      ProcessValue <- "MotorControl_Velocity_Velocity"
   Rectangle "Rectángulo_20" at 35,182 size 15x41
      Visibility <- "MotorControl_Velocity_Execute"
   Rectangle "Rectángulo_21" at 51,182 size 15x41
      Visibility <- "MotorControl_Velocity_Error"
   Rectangle "Rectángulo_22" at 19,182 size 15x41
      Visibility <- "MotorControl_Velocity_invelocity"
   TextField "Campo de texto_1" at 395,189 size 115x29; Text 'Velocidad / Velocity'
   IOField "Campo ES_7" at 524,13 size 142x40; FormatPattern s9999999999
      ProcessValue <- "2_PWMValve_Frecuency"
   TextField "Campo de texto_5" at 667,18 size 127x29; Text 'Frecuencia / Frequency'
   IOField "Campo ES_8" at 523,67 size 145x40; FormatPattern s99999
      ProcessValue <- "2_PWMValve_Duty_Cycle"
   TextField "Campo de texto_10" at 675,72 size 94x29; Text 'Trabajo / Duty'
   Rectangle "Rectángulo_18" at 575,117 size 15x41
      Visibility <- "2_PWMValve_Enable"
   Rectangle "Rectángulo_19" at 591,117 size 15x41
      Visibility <- "2_PWMValve_Busy"
   Rectangle "Rectángulo_38" at 559,117 size 15x41
      Visibility <- "2_PWMValve_Status"
   Button "Botón_9" at 610,184 size 145x40; TextOff 'MEM VELOC. / MEM SPEED'
      on Press: function_b14e0dd5("MotorControl_Velocity_Current", 0)
   TextField "Campo de texto_9" at 524,445 size 101x27; Text 'BATERIA / BATTERY'
   IOField "Campo ES_14" at 619,442 size 89x35; FormatPattern 99.9; Unit  Vdc
      ProcessValue <- "DataValues_BatteryVoltage"
   Button "Botón_14" at 534,442 size 35x35; TextOff 'M'
      on Press: ActivateScreen("Start", 0)
   IOField "Campo ES_15" at 711,442 size 82x35; FormatPattern 999.9; Unit  %
      ProcessValue <- "DataValues_BatteryCapacity"
   Button "Botón_18" at 582,442 size 35x35; TextOff 'M'
      on Press: ActivateScreen("Motor", 0)
   Button "Botón_1" at 7,442 size 80x35; TextOff 'GRAFICOS / GRAPHICS'
      on Press: ActivateScreen("Graphics", 0)
   Button "Botón_3" at 92,442 size 80x35; TextOff 'DATOS / DATA'
      on Press: ActivateScreen("Parameters", 0)
   Button "Botón_4" at 347,442 size 80x35; TextOff 'MANUALES / MANUALS'
      on Press: ActivateScreen("UserManual", 0)
   Button "Botón_5" at 432,442 size 80x35; TextOff 'ALARMAS / ALARMS'
      on Press: ActivateScreen("Alarms", 0)
   Button "Botón_12" at 177,442 size 80x35; TextOff 'PACIENTE / PATIENT'
      on Press: function_efd93a16("PatientData", 0, 0, 1, -1, 1)
   Button "Botón_19" at 262,442 size 80x35; TextOff 'RPM / BPM'
      on Press: function_efd93a16("RespirationRatios", 0, 0, 1, -1, 1)
   IOField "Campo ES_9" at 243,57 size 142x40; FormatPattern 9999
      ProcessValue <- "TurnAxis_Position"
   TextField "Campo de texto_11" at 396,62 size 100x29; Text 'Posición / Position'

PopupScreen "ControlMode" 600x300
   TextField "Campo de texto_2" at 107,59 size 238x39; Text 'Selección TIPO / Select TYPE'
   TextField "Campo de texto_1" at 204,5 size 192x30; Text 'MODO CONTROL / CONTROL MODE'
   SymbolicIOField "Campo ES simbólico_1" at 114,119 size 360x47; TextOff '0'; TextOn '1'; TextList "ControlMode"
      ProcessValue <- "OperatingParameters_ControlMode"
   Button "Botón_6" at 429,255 size 146x32; TextOff 'Salida / Exit'
      on Click: function_efd93a16("ControlMode", 0, 0, 0, -1, 1)
   IOField "Campo ES_8" at 23,255 size 242x32; FormatPattern 99999999999999999999
      ProcessValue <- "DateTime_LocalDateOut"

PopupScreen "Alarm" 400x300
   TextField "Campo de texto_1" at 41,95 size 315x91; Text 'ALARMA / ALARM'

PopupScreen "PatientData" 600x300
   TextField "Campo de texto_2" at 167,65 size 60x29; Text 'Sexo / Sex'
   TextField "Campo de texto_3" at 264,113 size 166x29; Text 'Volumen Tidal / Tidal Volume'
   TextField "Campo de texto_10" at 53,113 size 80x29; Text 'Altura / Height'
   IOField "Campo ES_6" at 138,110 size 110x35; FormatPattern 9.99; Unit m
      ProcessValue <- "PatientData_PatientHeight"
   IOField "Campo ES_11" at 432,110 size 110x35; FormatPattern 999.9; Unit ml
      ProcessValue <- "PatientData_TidalVolume"
   TextField "Campo de texto_1" at 198,8 size 204x30; Text 'DATOS PACIENTE / PATIENT DATA'
   SymbolicIOField "Campo ES simbólico_1" at 227,61 size 233x37; TextOn '1'; TextOff '0'; TextList "PatientSex"
      ProcessValue <- "PatientData_PatientType"
   Button "Botón_6" at 429,255 size 146x32; TextOff 'Salida / Exit'
      on Click: function_efd93a16("PatientData", 0, 0, 0, -1, 1)
   IOField "Campo ES_8" at 23,255 size 242x32; FormatPattern 99999999999999999999
      ProcessValue <- "DateTime_LocalDateOut"

PopupScreen "Pip" 600x300
   TextField "Campo de texto_2" at 242,90 size 46x29; Text 'PIP'
   IOField "Campo ES_8" at 389,87 size 75x35; Authorization "Operación"; FormatPattern 999
      ProcessValue <- "DataValues_PipValue"
   IOField "Campo ES_2" at 290,87 size 75x35; FormatPattern 999
      ProcessValue <- "OperatingParameters_PipMax"
   IOField "Campo ES_3" at 44,87 size 75x35; FormatPattern 999
      ProcessValue <- "OperatingParameters_PipSetpoint"
      Visibility <- "OperatingParameters_ControlMode"
   TextField "Campo de texto_5" at 34,44 size 128x29; Text 'CONSIGNA / SETPOINT'
   TextField "Campo de texto_6" at 300,44 size 55x29; Text 'MAX'
   TextField "Campo de texto_7" at 388,44 size 81x29; Text 'VALOR / VALUE'
   TextField "Campo de texto_8" at 496,44 size 56x29; Text 'MIN'
   IOField "Campo ES_7" at 485,87 size 75x35; FormatPattern 999
      ProcessValue <- "OperatingParameters_PipMin"
   IOField "Campo ES_1" at 290,141 size 75x35; FormatPattern 999
      ProcessValue <- "ProcessData_PpipSetpointAlarmHI"
   IOField "Campo ES_4" at 485,141 size 75x35; FormatPattern 999
      ProcessValue <- "ProcessData_PipSetpointAlarmLOW"
   IOField "Campo ES_5" at 290,195 size 75x35; FormatPattern 999
      ProcessValue <- "ProcessData_PipSetpointPreAlarmHI"
   IOField "Campo ES_6" at 485,195 size 75x35; FormatPattern 999
      ProcessValue <- "ProcessData_PipSetpointPreAlarmLOW"
   TextField "Campo de texto_1" at 155,144 size 134x29; Text 'PIP Alarma / PIP Alarm'
   TextField "Campo de texto_3" at 131,196 size 158x29; Text 'PIP PreAlarm'
   TextField "Campo de texto_4" at 187,8 size 226x30; Text 'PARAMETROS PEEP / PIP PARAMETERS'
   Button "Botón_6" at 429,255 size 146x32; TextOff 'Salida / Exit'
      on Click: function_efd93a16("Pip", 0, 0, 0, -1, 1)
   IOField "Campo ES_9" at 23,255 size 242x32; FormatPattern 99999999999999999999
      ProcessValue <- "DateTime_LocalDateOut"
   GraphicIOField "PlotLight_Round_GN_1" at 369,105 size 17x17; PictureOff "gris"; PictureOn "amarillo"
      ProcessValue <- "AlarmsRaw_PipDisplayPreAlarmHI"
   GraphicIOField "PlotLight_Round_GN_2" at 466,105 size 17x17; PictureOff "gris"; PictureOn "rojo"
      ProcessValue <- "AlarmsRaw_PipDisplayAlarmLOW"
   GraphicIOField "PlotLight_Round_GN_3" at 369,87 size 17x17; PictureOff "gris"; PictureOn "rojo"
      ProcessValue <- "AlarmsRaw_PipDisplayAlarmHI"
   GraphicIOField "PlotLight_Round_GN_4" at 466,87 size 17x17; PictureOff "gris"; PictureOn "amarillo"
      ProcessValue <- "AlarmsRaw_PipDisplayPreAlarmLOW"

PopupScreen "Plateau" 600x300
   TextField "Campo de texto_2" at 193,89 size 92x29; Text 'Plateau'
   IOField "Campo ES_8" at 389,87 size 75x35; Authorization "Operación"; FormatPattern 999
      ProcessValue <- "DataValues_PlateauValue"
   IOField "Campo ES_2" at 290,87 size 75x35; FormatPattern 999
      ProcessValue <- "OperatingParameters_PlateauMax"
   TextField "Campo de texto_5" at 34,44 size 128x29; Text 'CONSIGNA / SETPOINT'
   TextField "Campo de texto_6" at 300,44 size 55x29; Text 'MAX'
   TextField "Campo de texto_7" at 387,44 size 81x29; Text 'VALOR / VALUE'
   TextField "Campo de texto_8" at 496,44 size 56x29; Text 'MIN'
   IOField "Campo ES_7" at 485,87 size 75x35; FormatPattern 999
      ProcessValue <- "OperatingParameters_PlateauMin"
   IOField "Campo ES_1" at 290,141 size 75x35; FormatPattern 999
      ProcessValue <- "ProcessData_PlateauSetpointAlarmHI"
   IOField "Campo ES_4" at 485,141 size 75x35; FormatPattern 999
      ProcessValue <- "ProcessData_PlateaukSetpointAlarmLOW"
   IOField "Campo ES_5" at 290,195 size 75x35; FormatPattern 999
      ProcessValue <- "ProcessData_PlateauSetpointPreAlarmHI"
   IOField "Campo ES_6" at 485,195 size 75x35; FormatPattern 999
      ProcessValue <- "ProcessData_PlateauSetpointPreAlarmLOW"
   TextField "Campo de texto_1" at 119,144 size 166x29; Text 'Plateau Alarm'
   TextField "Campo de texto_3" at 81,198 size 204x29; Text 'Plateau PreAlarm'
   TextField "Campo de texto_4" at 165,7 size 271x30; Text 'PARAMETROS PLATEAU / PLATEAU PARAMETERS'
   Button "Botón_6" at 429,255 size 146x32; TextOff 'Salida / Exit'
      on Click: function_efd93a16("Plateau", 0, 0, 0, -1, 1)
   IOField "Campo ES_9" at 23,255 size 242x32; FormatPattern 99999999999999999999
      ProcessValue <- "DateTime_LocalDateOut"
   GraphicIOField "PlotLight_Round_GN_1" at 368,106 size 17x17; PictureOff "gris"; PictureOn "amarillo"
      ProcessValue <- "AlarmsRaw_PlateauDisplayPreAlarmHI"
   GraphicIOField "PlotLight_Round_GN_7" at 465,106 size 17x17; PictureOff "gris"; PictureOn "rojo"
      ProcessValue <- "AlarmsRaw_PlateauDisplayAlarmLOW"
   GraphicIOField "PlotLight_Round_GN_13" at 368,88 size 17x17; PictureOff "gris"; PictureOn "rojo"
      ProcessValue <- "AlarmsRaw_PlateauDisplayAlarmHI"
   GraphicIOField "PlotLight_Round_GN_19" at 465,88 size 17x17; PictureOff "gris"; PictureOn "amarillo"
      ProcessValue <- "AlarmsRaw_PlateauDisplayPreAlarmLOW"

PopupScreen "Peep" 600x300
   TextField "Campo de texto_2" at 225,88 size 60x29; Text 'Peep'
   IOField "Campo ES_8" at 391,87 size 75x35; Authorization "Operación"; FormatPattern 999
      ProcessValue <- "DataValues_PeepValue"
   IOField "Campo ES_2" at 290,87 size 75x35; FormatPattern 999
      ProcessValue <- "OperatingParameters_PeepMax"
   IOField "Campo ES_3" at 44,87 size 75x35; FormatPattern 999
      ProcessValue <- "OperatingParameters_PeepSetpoint"
      Visibility <- "OperatingParameters_ControlMode"
   TextField "Campo de texto_5" at 34,44 size 128x29; Text 'CONSIGNA / SETPOINT'
   TextField "Campo de texto_6" at 300,44 size 55x29; Text 'MAX'
   TextField "Campo de texto_7" at 389,44 size 81x29; Text 'VALOR / VALUE'
   TextField "Campo de texto_8" at 496,44 size 56x29; Text 'MIN'
   IOField "Campo ES_7" at 485,87 size 75x35; FormatPattern 999
      ProcessValue <- "OperatingParameters_PeepMin"
   IOField "Campo ES_1" at 290,141 size 75x35; FormatPattern 999
      ProcessValue <- "ProcessData_PeepSetpointAlarmHI"
   IOField "Campo ES_4" at 485,141 size 75x35; FormatPattern 999
      ProcessValue <- "ProcessData_PeepSetpointAlarmLOW"
   IOField "Campo ES_5" at 290,195 size 75x35; FormatPattern 999
      ProcessValue <- "ProcessData_PeepSetpointPreAlarmHI"
   IOField "Campo ES_6" at 485,195 size 75x35; FormatPattern 999
      ProcessValue <- "ProcessData_PeepSetpointPreAlarmLOW"
   TextField "Campo de texto_1" at 141,143 size 148x29; Text 'Peep Alarma / Peep Alarm'
   TextField "Campo de texto_3" at 103,197 size 186x29; Text 'Peep PreAlarma / Peep PreAlarm'
   TextField "Campo de texto_4" at 187,8 size 226x30; Text 'PARAMETROS PEEP / PEEP PARAMETERS'
   Button "Botón_6" at 429,255 size 146x32; TextOff 'Salida / Exit'
      on Click: function_efd93a16("Peep", 0, 0, 0, -1, 1)
   IOField "Campo ES_9" at 23,255 size 242x32; FormatPattern 99999999999999999999
      ProcessValue <- "DateTime_LocalDateOut"
   GraphicIOField "PlotLight_Round_GN_2" at 370,104 size 17x17; PictureOff "gris"; PictureOn "amarillo"
      ProcessValue <- "AlarmsRaw_PeepDisplayPreAlarmHI"
   GraphicIOField "PlotLight_Round_GN_8" at 467,104 size 17x17; PictureOff "gris"; PictureOn "rojo"
      ProcessValue <- "AlarmsRaw_PeepDisplayAlarmLOW"
   GraphicIOField "PlotLight_Round_GN_14" at 370,86 size 17x17; PictureOff "gris"; PictureOn "rojo"
      ProcessValue <- "AlarmsRaw_PeepDisplayAlarmHI"
   GraphicIOField "PlotLight_Round_GN_20" at 467,86 size 17x17; PictureOff "gris"; PictureOn "amarillo"
      ProcessValue <- "AlarmsRaw_PeepDisplayPreAlarmLOW"

PopupScreen "Frecuency" 600x300
   TextField "Campo de texto_2" at 161,89 size 127x29; Text 'Frecuencia / Frequency'
   IOField "Campo ES_8" at 388,87 size 75x35; Authorization "Operación"; FormatPattern 999
      ProcessValue <- "DataValues_FrequencyValue"
   IOField "Campo ES_2" at 290,87 size 75x35; FormatPattern 999
      ProcessValue <- "OperatingParameters_FrequencyMax"
   IOField "Campo ES_3" at 44,87 size 75x35; FormatPattern 999
      ProcessValue <- "OperatingParameters_FrequencySetpoint"
   TextField "Campo de texto_5" at 34,44 size 128x29; Text 'CONSIGNA / SETPOINT'
   TextField "Campo de texto_6" at 300,44 size 55x29; Text 'MAX'
   TextField "Campo de texto_7" at 387,44 size 81x29; Text 'VALOR / VALUE'
   TextField "Campo de texto_8" at 496,44 size 56x29; Text 'MIN'
   IOField "Campo ES_7" at 485,87 size 75x35; FormatPattern 999
      ProcessValue <- "OperatingParameters_FrequencyMin"
   IOField "Campo ES_1" at 290,141 size 75x35; FormatPattern 999
      ProcessValue <- "ProcessData_FrequencySetpointAlarmHI"
   IOField "Campo ES_4" at 485,141 size 75x35; FormatPattern 999
      ProcessValue <- "ProcessData_FrequencySetpointAlarmLOW"
   IOField "Campo ES_5" at 290,195 size 75x35; FormatPattern 999
      ProcessValue <- "ProcessData_FrequencySetpointPreAlarmHI"
   IOField "Campo ES_6" at 485,195 size 75x35; FormatPattern 999
      ProcessValue <- "ProcessData_FrequencySetpointPreAlarmLOW"
   TextField "Campo de texto_1" at 73,144 size 215x29; Text 'Frecuencia Alarma / Frequency Alarm'
   TextField "Campo de texto_3" at 56,197 size 233x29; Text 'FrecuenciaPreAlarm / Frequency PreAlarm'
   TextField "Campo de texto_4" at 143,5 size 315x30; Text 'PARAMETROS FRECUENCIA / FREQUENCY PARAMETERS'
   Button "Botón_6" at 429,255 size 146x32; TextOff 'Salida / Exit'
      on Click: function_efd93a16("Frecuency", 0, 0, 0, -1, 1)
   IOField "Campo ES_9" at 23,255 size 242x32; FormatPattern 99999999999999999999
      ProcessValue <- "DateTime_LocalDateOut"
   GraphicIOField "PlotLight_Round_GN_3" at 369,105 size 17x17; PictureOff "gris"; PictureOn "amarillo"
      ProcessValue <- "AlarmsRaw_FrequencyDisplayPreAlarmHI"
   GraphicIOField "PlotLight_Round_GN_9" at 466,105 size 17x17; PictureOff "gris"; PictureOn "rojo"
      ProcessValue <- "AlarmsRaw_FrequencyDisplayAlarmLOW"
   GraphicIOField "PlotLight_Round_GN_15" at 369,87 size 17x17; PictureOff "gris"; PictureOn "rojo"
      ProcessValue <- "AlarmsRaw_FrequencyDisplayAlarmHI"
   GraphicIOField "PlotLight_Round_GN_21" at 466,87 size 17x17; PictureOff "gris"; PictureOn "amarillo"
      ProcessValue <- "AlarmsRaw_FrequencyDisplayPreAlarmLOW"

PopupScreen "TidalVolume" 600x300
   TextField "Campo de texto_2" at 123,90 size 166x29; Text 'Volumen Tidal / Tidal Volume'
   IOField "Campo ES_8" at 391,87 size 75x35; Authorization "Operación"; FormatPattern 999
      ProcessValue <- "DataValues_TidalVolumeValue"
   IOField "Campo ES_2" at 290,87 size 75x35; FormatPattern 999
      ProcessValue <- "OperatingParameters_TidalVolumenMax"
   IOField "Campo ES_3" at 44,87 size 75x35; FormatPattern 999
      ProcessValue <- "OperatingParameters_TidalVolumenSetpoint"
      Visibility <- "OperatingParameters_ControlMode"
   TextField "Campo de texto_5" at 34,44 size 128x29; Text 'CONSIGNA / SETPOINT'
   TextField "Campo de texto_6" at 300,44 size 55x29; Text 'MAX'
   TextField "Campo de texto_7" at 391,44 size 81x29; Text 'VALOR / VALUE'
   TextField "Campo de texto_8" at 496,44 size 56x29; Text 'MIN'
   IOField "Campo ES_7" at 485,87 size 75x35; FormatPattern 999
      ProcessValue <- "OperatingParameters_TidalVolumenMin"
   IOField "Campo ES_1" at 290,141 size 75x35; FormatPattern 999
      ProcessValue <- "ProcessData_TidalVolumeSetpointAlarmHI"
   IOField "Campo ES_4" at 485,141 size 75x35; FormatPattern 999
      ProcessValue <- "ProcessData_TidalVolumeSetpointAlarmLOW"
   IOField "Campo ES_5" at 290,195 size 75x35; FormatPattern 999
      ProcessValue <- "ProcessData_TidalVolumeSetpointPreAlarmHI"
   IOField "Campo ES_6" at 485,195 size 75x35; FormatPattern 999
      ProcessValue <- "ProcessData_TidalVolumeSetpointPreAlarmLOW"
   TextField "Campo de texto_1" at 35,143 size 254x29; Text 'Alarma Volumen Tidal / Tidal Volume Alarm'
   TextField "Campo de texto_3" at 0,197 size 290x29; Text 'PreAlarma volumen Tidal / Tidal Volume PreAlarm'
   TextField "Campo de texto_4" at 121,8 size 358x30; Text 'PARAMETROS VOLUMEN TIDAL / TIDAL VOLUME PARAMETERS'
   Button "Botón_6" at 429,255 size 146x32; TextOff 'Salida / Exit'
      on Click: function_efd93a16("TidalVolume", 0, 0, 0, -1, 1)
   IOField "Campo ES_9" at 23,255 size 242x32; FormatPattern 99999999999999999999
      ProcessValue <- "DateTime_LocalDateOut"
   GraphicIOField "PlotLight_Round_GN_4" at 370,105 size 17x17; PictureOff "gris"; PictureOn "amarillo"
      ProcessValue <- "AlarmsRaw_TidalVolumeDisplayPreAlarmHI"
   GraphicIOField "PlotLight_Round_GN_10" at 467,105 size 17x17; PictureOff "gris"; PictureOn "rojo"
      ProcessValue <- "AlarmsRaw_TidalVolumeDisplayAlarmLOW"
   GraphicIOField "PlotLight_Round_GN_16" at 370,87 size 17x17; PictureOff "gris"; PictureOn "rojo"
      ProcessValue <- "AlarmsRaw_TidalVolumeDisplayAlarmHI"
   GraphicIOField "PlotLight_Round_GN_22" at 467,87 size 17x17; PictureOff "gris"; PictureOn "amarillo"
      ProcessValue <- "AlarmsRaw_TidalVolumeDisplayPreAlarmLOW"

PopupScreen "VolumeMinute" 600x300
   TextField "Campo de texto_2" at 114,90 size 174x29; Text 'Vol. Minute / Minute Volume'
   IOField "Campo ES_8" at 388,87 size 75x35; Authorization "Operación"; FormatPattern 999
      ProcessValue <- "DataValues_MinumValue"
   IOField "Campo ES_2" at 290,87 size 75x35; FormatPattern 999
      ProcessValue <- "OperatingParameters_MinimumVolumeMax"
   IOField "Campo ES_3" at 44,87 size 75x35; FormatPattern 999
      Visibility <- "OperatingParameters_ControlMode"
      ProcessValue <- "OperatingParameters_MinimumVolumeSetpoint"
   TextField "Campo de texto_5" at 34,44 size 128x29; Text 'CONSIGNA / SETPOINT'
   TextField "Campo de texto_6" at 300,44 size 55x29; Text 'MAX'
   TextField "Campo de texto_7" at 390,44 size 81x29; Text 'VALOR / VALUE'
   TextField "Campo de texto_8" at 496,44 size 56x29; Text 'MIN'
   IOField "Campo ES_7" at 485,87 size 75x35; FormatPattern 999
      ProcessValue <- "OperatingParameters_MinimumVolumeMin"
   IOField "Campo ES_1" at 290,141 size 75x35; FormatPattern 999
      ProcessValue <- "ProcessData_VolumeMinSetpointAlarmHI"
   IOField "Campo ES_4" at 485,141 size 75x35; FormatPattern 999
      ProcessValue <- "ProcessData_VolumeMinSetpointPreAlarmLOW"
   IOField "Campo ES_5" at 290,195 size 75x35; FormatPattern 999
      ProcessValue <- "ProcessData_VolumeMinSetpointPreAlarmHI"
   IOField "Campo ES_6" at 485,195 size 75x35; FormatPattern 999
      ProcessValue <- "ProcessData_VolumeMinSetpointAlarmLOW"
   TextField "Campo de texto_1" at 20,143 size 269x29; Text 'Volumen/Minuto Alarm / Volume/Minute Alarm'
   TextField "Campo de texto_3" at 12,198 size 277x29; Text 'Volumen/Min. PreAlarm / Volume/Min. PreAlarm'
   TextField "Campo de texto_4" at 105,5 size 390x30; Text 'PARAMETROS VOLUMEN/MINUTO / VOLUME/MINUTE PARAMETERS'
   Button "Botón_6" at 429,255 size 146x32; TextOff 'Salida / Exit'
      on Click: function_efd93a16("VolumeMinute", 0, 0, 0, -1, 1)
   IOField "Campo ES_9" at 23,255 size 242x32; FormatPattern 99999999999999999999
      ProcessValue <- "DateTime_LocalDateOut"
   GraphicIOField "PlotLight_Round_GN_5" at 368,87 size 17x17; PictureOff "gris"; PictureOn "rojo"
      ProcessValue <- "AlarmsRaw_VolumeMinuteDisplayAlarmHI"
   GraphicIOField "PlotLight_Round_GN_11" at 465,105 size 17x17; PictureOff "gris"; PictureOn "rojo"
      ProcessValue <- "AlarmsRaw_VolumeMinuteDisplayAlarmLOW"
   GraphicIOField "PlotLight_Round_GN_17" at 368,105 size 17x17; PictureOff "gris"; PictureOn "amarillo"
      ProcessValue <- "AlarmsRaw_VolumeMinuteDisplayPreAlarmHI"
   GraphicIOField "PlotLight_Round_GN_23" at 465,87 size 17x17; PictureOff "gris"; PictureOn "amarillo"
      ProcessValue <- "AlarmsRaw_VolumeMinuteDisplayPreAlarmLOW"

PopupScreen "Trigger" 600x300
   TextField "Campo de texto_2" at 199,88 size 87x29; Text 'Trigger'
   IOField "Campo ES_8" at 388,87 size 75x35; Authorization "Operación"; FormatPattern 999
      ProcessValue <- "DataValues_Trigger"
   IOField "Campo ES_2" at 290,87 size 75x35; FormatPattern 999
      ProcessValue <- "OperatingParameters_TriggerMax"
   IOField "Campo ES_3" at 44,87 size 75x35; FormatPattern 999
      ProcessValue <- "OperatingParameters_TriggerSetpoint"
   TextField "Campo de texto_5" at 34,44 size 128x29; Text 'CONSIGNA / SETPOINT'
   TextField "Campo de texto_6" at 300,44 size 55x29; Text 'MAX'
   TextField "Campo de texto_7" at 387,44 size 81x29; Text 'VALOR / VALUE'
   TextField "Campo de texto_8" at 496,44 size 56x29; Text 'MIN'
   IOField "Campo ES_7" at 485,87 size 75x35; FormatPattern 999
      ProcessValue <- "OperatingParameters_TriggerMin"
   IOField "Campo ES_1" at 290,141 size 75x35; FormatPattern 999
      ProcessValue <- "ProcessData_TriggerVolumeSetpointAlarmHI"
   IOField "Campo ES_4" at 485,141 size 75x35; FormatPattern 999
      ProcessValue <- "ProcessData_TriggerVolumeSetpointAlarmLOW"
   IOField "Campo ES_5" at 290,195 size 75x35; FormatPattern 999
      ProcessValue <- "ProcessData_TriggeVolumeSetpointPreAlarmHI"
   IOField "Campo ES_6" at 485,195 size 75x35; FormatPattern 999
      ProcessValue <- "ProcessData_TriggerVolumeSetpointPreAlarmLOW"
   TextField "Campo de texto_1" at 125,143 size 161x29; Text 'Trigger Alarm'
   TextField "Campo de texto_3" at 87,197 size 199x29; Text 'Trigger PreAlarm'
   TextField "Campo de texto_4" at 164,8 size 273x30; Text 'PARAMETROS TRIGGER / TRIGGER PARAMETERS'
   Button "Botón_6" at 429,255 size 146x32; TextOff 'Salida / Exit'
      on Click: function_efd93a16("Trigger", 0, 0, 0, -1, 1)
   Button "Botón_7" at 396,141 size 61x35; TextOff 'Trigger'
      Visibility <- "Clock_1Hz"
   TextField "Campo de texto_9" at 396,196 size 61x35; Text 'OFF'
      Visibility <- "OperatingParameters_Trigger"
   TextField "Campo de texto_10" at 396,196 size 61x35; Text 'ON'
      Visibility <- "OperatingParameters_Trigger"
   Button "Botón_1" at 396,196 size 61x35; TextOn 'ON'; TextOff 'Text'
      on Click: InvertBit("OperatingParameters_Trigger")
      Appearance <- "OperatingParameters_Trigger"
   IOField "Campo ES_9" at 23,255 size 242x32; FormatPattern 99999999999999999999
      ProcessValue <- "DateTime_LocalDateOut"
   GraphicIOField "PlotLight_Round_GN_4" at 370,105 size 17x17; PictureOn "amarillo"; PictureOff "gris"
      ProcessValue <- "AlarmsRaw_TriggerDisplayPreAlarmHI"
   GraphicIOField "PlotLight_Round_GN_10" at 467,105 size 17x17; PictureOn "rojo"; PictureOff "gris"
      ProcessValue <- "AlarmsRaw_TriggerDisplayAlarmLOW"
   GraphicIOField "PlotLight_Round_GN_16" at 370,87 size 17x17; PictureOn "rojo"; PictureOff "gris"
      ProcessValue <- "AlarmsRaw_TriggerDisplayAlarmHI"
   GraphicIOField "PlotLight_Round_GN_22" at 467,87 size 17x17; PictureOn "amarillo"; PictureOff "gris"
      ProcessValue <- "AlarmsRaw_TriggerDisplayPreAlarmLOW"

PopupScreen "Enviroment" 600x300
   TextField "Campo de texto_2" at 30,82 size 124x29; Text 'Humidif. / Humidifier'
   IOField "Campo ES_3" at 246,192 size 75x35; FormatPattern 999
      ProcessValue <- "OperatingParameters_O2Setpoint"
   TextField "Campo de texto_4" at 140,5 size 320x30; Text 'PARAMETROS ENTORNO / ENVIROMENT PARAMETERS'
   Button "Botón_6" at 429,255 size 146x32; TextOff 'Salida / Exit'
      on Click: function_efd93a16("Enviroment", 0, 0, 0, -1, 1)
   Button "Botón_7" at 429,79 size 61x35; TextOff 'Hr'
      Visibility <- "Clock_1Hz"
   TextField "Campo de texto_9" at 502,79 size 61x35; Text 'OFF'
      Visibility <- "OperatingParameters_Trigger"
   TextField "Campo de texto_10" at 502,79 size 61x35; Text 'ON'
      Visibility <- "OperatingParameters_Trigger"
   Button "Botón_1" at 506,79 size 61x35; TextOn 'ON'; TextOff 'Text'
      on Click: InvertBit("OperatingParameters_Trigger")
      Appearance <- "OperatingParameters_Trigger"
   IOField "Campo ES_5" at 330,80 size 89x35; FormatPattern 9999999
      ProcessValue <- "OperatingParameters_HumidifiertElap"
   IOField "Campo ES_1" at 237,80 size 89x35; FormatPattern 9999999
      ProcessValue <- "OperatingParameters_HumidifierTimer"
   TextField "Campo de texto_1" at 38,196 size 142x29; Text 'Presión O2 / O2 Pressure'
   Button "Botón_2" at 429,192 size 61x35; TextOff 'O2'
      Visibility <- "Clock_1Hz"
   TextField "Campo de texto_3" at 502,192 size 61x35; Text 'OFF'
      Visibility <- "OperatingParameters_O2"
   TextField "Campo de texto_5" at 502,192 size 61x35; Text 'ON'
      Visibility <- "OperatingParameters_O2"
   Button "Botón_3" at 506,192 size 61x35; TextOn 'ON'; TextOff 'Text'
      on Click: InvertBit("OperatingParameters_O2")
      Appearance <- "OperatingParameters_Trigger"
   TextField "Campo de texto_6" at 502,47 size 67x29; Text 'Modo / Mode'
   TextField "Campo de texto_7" at 418,47 size 83x29; Text 'Estado / State'
   TextField "Campo de texto_8" at 327,47 size 93x29; Text 'Trasn. / Elapsed'
   TextField "Campo de texto_11" at 246,48 size 75x29; Text 'Temp. / Timer'
   TextField "Campo de texto_12" at 38,156 size 143x29; Text 'Presión Aire / Air Pressure'
   Button "Botón_4" at 429,152 size 61x35; TextOff 'Aire / Air'
      Visibility <- "Clock_1Hz"
   TextField "Campo de texto_13" at 502,153 size 61x35; Text 'OFF'
      Visibility <- "OperatingParameters_Air"
   TextField "Campo de texto_14" at 502,153 size 61x35; Text 'ON'
      Visibility <- "OperatingParameters_Air"
   Button "Botón_5" at 506,153 size 61x35; TextOn 'ON'; TextOff 'Text'
      on Click: InvertBit("OperatingParameters_Air")
      Appearance <- "OperatingParameters_Trigger"
   IOField "Campo ES_2" at 336,192 size 75x35; FormatPattern 999
      ProcessValue <- "DataValues_O2Pressure"
   IOField "Campo ES_4" at 246,153 size 75x35; FormatPattern 999
      ProcessValue <- "OperatingParameters_AirSetpoint"
   IOField "Campo ES_6" at 336,153 size 75x35; FormatPattern 999
      ProcessValue <- "DataValues_AirPressure"
   TextField "Campo de texto_15" at 340,122 size 68x29; Text 'Valor / Value'
   TextField "Campo de texto_16" at 234,123 size 109x29; Text 'Consigna / Setpoint'
   IOField "Campo ES_7" at 144,80 size 89x35; FormatPattern 9999999
      ProcessValue <- "OperatingParameters_HumidifiertDuration"
   TextField "Campo de texto_17" at 156,48 size 67x29; Text 'Pulso / Pulse'
   IOField "Campo ES_8" at 23,255 size 242x32; FormatPattern 99999999999999999999
      ProcessValue <- "DateTime_LocalDateOut"

